// TIA Portal project "YDSLK_HMI_2023-05-10_08-26_V3_00T" (V15.1) (continued)
   "ST_HMI_Var_HMI_r64_DingZi_Zouche_ratio_KongDing_65_1" : LReal = PLC ST_HMI_Var.HMI_r64_DingZi_Zouche_ratio_KongDing_65_1 AT 10-30-00-01-00-21-84-00-4D-40, 1 s
   "ST_Calculation_Var_g_i16_Calculation_0_Status" : Int = PLC ST_Calculation_Var.g_i16_Calculation_0_Status AT 10-05-00-01-00-13-84-00-00-00, 1 s
   "ST_1TCP_g_myStructSend__lreal_20" : LReal = PLC ST_1TCP.g_myStructSend._lreal_20 AT 10-30-00-01-00-0D-84-01-30-40, 1 s
   "ST_1TCP_g_myStructSend__lreal_1" : LReal = PLC ST_1TCP.g_myStructSend._lreal_1 AT 10-30-00-01-00-0D-84-01-2B-80, 1 s
   "ST_HMI_Var_HMI_bo_ZouChe_Holding_Brake_Open" : Bool = PLC ST_HMI_Var.HMI_bo_ZouChe_Holding_Brake_Open AT 10-01-00-01-00-21-84-00-72-50, 1 s
   "ST_Real_Monitoring_HMI_r64_Real_QianShen_WuNian" : LReal = PLC ST_Real_Monitoring.HMI_r64_Real_QianShen_WuNian AT 10-30-00-01-00-2D-84-00-00-00, 1 s
   "ST_Real_Monitoring_HMI_r64Axis_ZouChe_Position_JiZhong_QianShen_Start" : LReal = PLC ST_Real_Monitoring.HMI_r64Axis_ZouChe_Position_JiZhong_QianShen_Start AT 10-30-00-01-00-2D-84-00-00-40, 1 s
   "ST_Real_Monitoring_HMI_r64_NianDu_JiZhong_QianShen_Start" : LReal = PLC ST_Real_Monitoring.HMI_r64_NianDu_JiZhong_QianShen_Start AT 10-30-00-01-00-2D-84-00-00-80, 1 s
   "ST_Real_Monitoring_HMI_r64Axis_ZouChe_Position_LuoLa_Stop" : LReal = PLC ST_Real_Monitoring.HMI_r64Axis_ZouChe_Position_LuoLa_Stop AT 10-30-00-01-00-2D-84-00-00-C0, 1 s
   "ST_Real_Monitoring_HMI_r64_NianDu_LuoLa_Stop" : LReal = PLC ST_Real_Monitoring.HMI_r64_NianDu_LuoLa_Stop AT 10-30-00-01-00-2D-84-00-01-00, 1 s
   "ST_Real_Monitoring_HMI_r64Axis_ZouChe_Position_YiNian_DaoDa" : LReal = PLC ST_Real_Monitoring.HMI_r64Axis_ZouChe_Position_YiNian_DaoDa AT 10-30-00-01-00-2D-84-00-01-40, 1 s
   "ST_Convert_ReadParameters_g_r64_SERVO_03_ZouChe_35_Motor_temperature_real" : LReal = PLC ST_Convert_ReadParameters.g_r64_SERVO_03_ZouChe_35_Motor_temperature_real AT 10-30-00-01-00-18-84-00-00-C0, 1 s
   "ST_Convert_ReadParameters_g_r64_SERVO_03_ZouChe_37_4_Power_unit_temperatures_Interior_of_power_unit_real" : LReal = PLC ST_Convert_ReadParameters.g_r64_SERVO_03_ZouChe_37_4_Power_unit_temperatures_Interior_of_power_unit_real AT 10-30-00-01-00-18-84-00-01-40, 1 s
   "ST_Convert_ReadParameters_g_r64_SERVO_04_ZhangLi_35_Motor_temperature_real" : LReal = PLC ST_Convert_ReadParameters.g_r64_SERVO_04_ZhangLi_35_Motor_temperature_real AT 10-30-00-01-00-18-84-00-03-00, 1 s
   "ST_Convert_ReadParameters_g_r64_SERVO_05_ChengXing_35_Motor_temperature_real" : LReal = PLC ST_Convert_ReadParameters.g_r64_SERVO_05_ChengXing_35_Motor_temperature_real AT 10-30-00-01-00-18-84-00-05-40, 1 s
   "ST_Convert_ReadParameters_g_r64_SERVO_06_GunTong_35_Motor_temperature_real" : LReal = PLC ST_Convert_ReadParameters.g_r64_SERVO_06_GunTong_35_Motor_temperature_real AT 10-30-00-01-00-18-84-00-07-80, 1 s
   "ST_Convert_ReadParameters_g_r64_SERVO_08_LuoLa_35_Motor_temperature_real" : LReal = PLC ST_Convert_ReadParameters.g_r64_SERVO_08_LuoLa_35_Motor_temperature_real AT 10-30-00-01-00-18-84-00-0C-00, 1 s
   "ST_Convert_ReadParameters_g_r64_SERVO_07_DingZi_35_Motor_temperature_real" : LReal = PLC ST_Convert_ReadParameters.g_r64_SERVO_07_DingZi_35_Motor_temperature_real AT 10-30-00-01-00-18-84-00-09-C0, 1 s
   "ST_Convert_ReadParameters_g_r64_SERVO_05_ChengXing_37_4_Power_unit_temperatures_Interior_of_power_unit_real" : LReal = PLC ST_Convert_ReadParameters.g_r64_SERVO_05_ChengXing_37_4_Power_unit_temperatures_Interior_of_power_unit_real AT 10-30-00-01-00-18-84-00-05-C0, 1 s
   "ST_Convert_ReadParameters_g_r64_SERVO_07_DingZi_37_4_Power_unit_temperatures_Interior_of_power_unit_real" : LReal = PLC ST_Convert_ReadParameters.g_r64_SERVO_07_DingZi_37_4_Power_unit_temperatures_Interior_of_power_unit_real AT 10-30-00-01-00-18-84-00-0A-40, 1 s
   "ST_Convert_ReadParameters_g_r64_SERVO_08_LuoLa_37_4_Power_unit_temperatures_Interior_of_power_unit_real" : LReal = PLC ST_Convert_ReadParameters.g_r64_SERVO_08_LuoLa_37_4_Power_unit_temperatures_Interior_of_power_unit_real AT 10-30-00-01-00-18-84-00-0C-80, 1 s

HMI tags "变量表_卷绕经验参数"
   "ST_Calculation_Var_1_ZhiShu_ARRAY_JR{3}" : LReal = PLC ST_Calculation_Var_1.ZhiShu_ARRAY_JR[3] AT 10-30-00-01-00-14-84-00-22-00, 1 s
   "ST_Calculation_Var_1_ZhiShu_ARRAY_JR{4}" : LReal = PLC ST_Calculation_Var_1.ZhiShu_ARRAY_JR[4] AT 10-30-00-01-00-14-84-00-22-40, 1 s
   "ST_Calculation_Var_1_ZhiShu_ARRAY_JR{5}" : LReal = PLC ST_Calculation_Var_1.ZhiShu_ARRAY_JR[5] AT 10-30-00-01-00-14-84-00-22-80, 1 s
   "ST_Calculation_Var_1_ZhiShu_ARRAY_JR{6}" : LReal = PLC ST_Calculation_Var_1.ZhiShu_ARRAY_JR[6] AT 10-30-00-01-00-14-84-00-22-C0, 1 s
   "ST_Calculation_Var_1_ZhiShu_ARRAY_JR{7}" : LReal = PLC ST_Calculation_Var_1.ZhiShu_ARRAY_JR[7] AT 10-30-00-01-00-14-84-00-23-00, 1 s
   "ST_Calculation_Var_1_ZhiShu_ARRAY_JR{8}" : LReal = PLC ST_Calculation_Var_1.ZhiShu_ARRAY_JR[8] AT 10-30-00-01-00-14-84-00-23-40, 1 s
   "ST_Calculation_Var_1_ZhiShu_ARRAY_JR{9}" : LReal = PLC ST_Calculation_Var_1.ZhiShu_ARRAY_JR[9] AT 10-30-00-01-00-14-84-00-23-80, 1 s
   "ST_Calculation_Var_1_ZhiShu_ARRAY_JR{10}" : LReal = PLC ST_Calculation_Var_1.ZhiShu_ARRAY_JR[10] AT 10-30-00-01-00-14-84-00-23-C0, 1 s
   "ST_Calculation_Var_1_ZhiShu_ARRAY_JR{11}" : LReal = PLC ST_Calculation_Var_1.ZhiShu_ARRAY_JR[11] AT 10-30-00-01-00-14-84-00-24-00, 1 s
   "ST_Calculation_Var_1_ZhiShu_ARRAY_JR{12}" : LReal = PLC ST_Calculation_Var_1.ZhiShu_ARRAY_JR[12] AT 10-30-00-01-00-14-84-00-24-40, 1 s
   "ST_Calculation_Var_1_ZhiShu_ARRAY_JR{13}" : LReal = PLC ST_Calculation_Var_1.ZhiShu_ARRAY_JR[13] AT 10-30-00-01-00-14-84-00-24-80, 1 s
   "ST_Calculation_Var_1_ZhiShu_ARRAY_JR{14}" : LReal = PLC ST_Calculation_Var_1.ZhiShu_ARRAY_JR[14] AT 10-30-00-01-00-14-84-00-24-C0, 1 s
   "ST_Calculation_Var_1_ZhiShu_ARRAY_JR{15}" : LReal = PLC ST_Calculation_Var_1.ZhiShu_ARRAY_JR[15] AT 10-30-00-01-00-14-84-00-25-00, 1 s
   "ST_Calculation_Var_1_ZhiShu_ARRAY_JR{16}" : LReal = PLC ST_Calculation_Var_1.ZhiShu_ARRAY_JR[16] AT 10-30-00-01-00-14-84-00-25-40, 1 s
   "ST_Calculation_Var_1_ZhiShu_ARRAY_JR{17}" : LReal = PLC ST_Calculation_Var_1.ZhiShu_ARRAY_JR[17] AT 10-30-00-01-00-14-84-00-25-80, 1 s
   "ST_Calculation_Var_1_ZhiShu_ARRAY_JR{18}" : LReal = PLC ST_Calculation_Var_1.ZhiShu_ARRAY_JR[18] AT 10-30-00-01-00-14-84-00-25-C0, 1 s
   "ST_Calculation_Var_1_ZhiShu_ARRAY_JR{19}" : LReal = PLC ST_Calculation_Var_1.ZhiShu_ARRAY_JR[19] AT 10-30-00-01-00-14-84-00-26-00, 1 s
   "ST_Calculation_Var_1_ZhiShu_ARRAY_JR{20}" : LReal = PLC ST_Calculation_Var_1.ZhiShu_ARRAY_JR[20] AT 10-30-00-01-00-14-84-00-26-40, 1 s
   "ST_Calculation_Var_1_ZhiShu_ARRAY_JR{21}" : LReal = PLC ST_Calculation_Var_1.ZhiShu_ARRAY_JR[21] AT 10-30-00-01-00-14-84-00-26-80, 1 s
   "ST_Calculation_Var_1_ZhiShu_ARRAY_JR{22}" : LReal = PLC ST_Calculation_Var_1.ZhiShu_ARRAY_JR[22] AT 10-30-00-01-00-14-84-00-26-C0, 1 s
   "ST_Calculation_Var_1_ZhiShu_ARRAY_JR{23}" : LReal = PLC ST_Calculation_Var_1.ZhiShu_ARRAY_JR[23] AT 10-30-00-01-00-14-84-00-27-00, 1 s
   "ST_Calculation_Var_1_ZhiShu_ARRAY_JR{24}" : LReal = PLC ST_Calculation_Var_1.ZhiShu_ARRAY_JR[24] AT 10-30-00-01-00-14-84-00-27-40, 1 s
   "ST_Calculation_Var_1_ZhiShu_ARRAY_JR{25}" : LReal = PLC ST_Calculation_Var_1.ZhiShu_ARRAY_JR[25] AT 10-30-00-01-00-14-84-00-27-80, 1 s
   "ST_Calculation_Var_1_ZhiShu_ARRAY_JR{26}" : LReal = PLC ST_Calculation_Var_1.ZhiShu_ARRAY_JR[26] AT 10-30-00-01-00-14-84-00-27-C0, 1 s
   "ST_Calculation_Var_1_ZhiShu_ARRAY_JR{27}" : LReal = PLC ST_Calculation_Var_1.ZhiShu_ARRAY_JR[27] AT 10-30-00-01-00-14-84-00-28-00, 1 s
   "ST_Calculation_Var_1_ZhiShu_ARRAY_JR{28}" : LReal = PLC ST_Calculation_Var_1.ZhiShu_ARRAY_JR[28] AT 10-30-00-01-00-14-84-00-28-40, 1 s
   "ST_Calculation_Var_1_ZhiShu_ARRAY_JR{29}" : LReal = PLC ST_Calculation_Var_1.ZhiShu_ARRAY_JR[29] AT 10-30-00-01-00-14-84-00-28-80, 1 s
   "ST_Calculation_Var_1_ZhiShu_ARRAY_JR{30}" : LReal = PLC ST_Calculation_Var_1.ZhiShu_ARRAY_JR[30] AT 10-30-00-01-00-14-84-00-28-C0, 1 s
   "ST_Calculation_Var_1_ZhiShu_ARRAY_JR{31}" : LReal = PLC ST_Calculation_Var_1.ZhiShu_ARRAY_JR[31] AT 10-30-00-01-00-14-84-00-29-00, 1 s
   "ST_Calculation_Var_1_ZhiShu_ARRAY_JR{32}" : LReal = PLC ST_Calculation_Var_1.ZhiShu_ARRAY_JR[32] AT 10-30-00-01-00-14-84-00-29-40, 1 s
   "ST_Calculation_Var_1_ZhiShu_ARRAY_JR{33}" : LReal = PLC ST_Calculation_Var_1.ZhiShu_ARRAY_JR[33] AT 10-30-00-01-00-14-84-00-29-80, 1 s
   "ST_Calculation_Var_1_ZhiShu_ARRAY_JR{34}" : LReal = PLC ST_Calculation_Var_1.ZhiShu_ARRAY_JR[34] AT 10-30-00-01-00-14-84-00-29-C0, 1 s
   "ST_Calculation_Var_1_ZhiShu_ARRAY_JR{35}" : LReal = PLC ST_Calculation_Var_1.ZhiShu_ARRAY_JR[35] AT 10-30-00-01-00-14-84-00-2A-00, 1 s
   "ST_Calculation_Var_1_ZhiShu_ARRAY_JR{36}" : LReal = PLC ST_Calculation_Var_1.ZhiShu_ARRAY_JR[36] AT 10-30-00-01-00-14-84-00-2A-40, 1 s
   "ST_Calculation_Var_1_ZhiShu_ARRAY_JR{37}" : LReal = PLC ST_Calculation_Var_1.ZhiShu_ARRAY_JR[37] AT 10-30-00-01-00-14-84-00-2A-80, 1 s
   "ST_Calculation_Var_1_ZhiShu_ARRAY_JR{38}" : LReal = PLC ST_Calculation_Var_1.ZhiShu_ARRAY_JR[38] AT 10-30-00-01-00-14-84-00-2A-C0, 1 s
   "ST_Calculation_Var_1_ZhiShu_ARRAY_JR{39}" : LReal = PLC ST_Calculation_Var_1.ZhiShu_ARRAY_JR[39] AT 10-30-00-01-00-14-84-00-2B-00, 1 s
   "ST_Calculation_Var_1_ZhiShu_ARRAY_JR{40}" : LReal = PLC ST_Calculation_Var_1.ZhiShu_ARRAY_JR[40] AT 10-30-00-01-00-14-84-00-2B-40, 1 s
   "ST_Calculation_Var_1_ZhiShu_ARRAY_JR{41}" : LReal = PLC ST_Calculation_Var_1.ZhiShu_ARRAY_JR[41] AT 10-30-00-01-00-14-84-00-2B-80, 1 s
   "ST_Calculation_Var_1_ZhiShu_ARRAY_JR{42}" : LReal = PLC ST_Calculation_Var_1.ZhiShu_ARRAY_JR[42] AT 10-30-00-01-00-14-84-00-2B-C0, 1 s
   "ST_Calculation_Var_1_ZhiShu_ARRAY_JR{43}" : LReal = PLC ST_Calculation_Var_1.ZhiShu_ARRAY_JR[43] AT 10-30-00-01-00-14-84-00-2C-00, 1 s
   "ST_Calculation_Var_1_ZhiShu_ARRAY_JR{44}" : LReal = PLC ST_Calculation_Var_1.ZhiShu_ARRAY_JR[44] AT 10-30-00-01-00-14-84-00-2C-40, 1 s
   "ST_Calculation_Var_1_ZhiShu_ARRAY_JR{45}" : LReal = PLC ST_Calculation_Var_1.ZhiShu_ARRAY_JR[45] AT 10-30-00-01-00-14-84-00-2C-80, 1 s
   "ST_Calculation_Var_1_ZhiShu_ARRAY_JR{46}" : LReal = PLC ST_Calculation_Var_1.ZhiShu_ARRAY_JR[46] AT 10-30-00-01-00-14-84-00-2C-C0, 1 s
   "ST_Calculation_Var_1_ZhiShu_ARRAY_JR{47}" : LReal = PLC ST_Calculation_Var_1.ZhiShu_ARRAY_JR[47] AT 10-30-00-01-00-14-84-00-2D-00, 1 s
   "ST_Calculation_Var_1_f1_n_delt_0_n_ARRAY_JR{3}" : LReal = PLC ST_Calculation_Var_1.f1_n_delt_0_n_ARRAY_JR[3] AT 10-30-00-01-00-14-84-00-2E-00, 1 s
   "ST_Calculation_Var_1_f1_n_delt_0_n_ARRAY_JR{4}" : LReal = PLC ST_Calculation_Var_1.f1_n_delt_0_n_ARRAY_JR[4] AT 10-30-00-01-00-14-84-00-2E-40, 1 s
   "ST_Calculation_Var_1_f1_n_delt_0_n_ARRAY_JR{5}" : LReal = PLC ST_Calculation_Var_1.f1_n_delt_0_n_ARRAY_JR[5] AT 10-30-00-01-00-14-84-00-2E-80, 1 s
   "ST_Calculation_Var_1_f1_n_delt_0_n_ARRAY_JR{6}" : LReal = PLC ST_Calculation_Var_1.f1_n_delt_0_n_ARRAY_JR[6] AT 10-30-00-01-00-14-84-00-2E-C0, 1 s
   "ST_Calculation_Var_1_f1_n_delt_0_n_ARRAY_JR{7}" : LReal = PLC ST_Calculation_Var_1.f1_n_delt_0_n_ARRAY_JR[7] AT 10-30-00-01-00-14-84-00-2F-00, 1 s
   "ST_Calculation_Var_1_f1_n_delt_0_n_ARRAY_JR{8}" : LReal = PLC ST_Calculation_Var_1.f1_n_delt_0_n_ARRAY_JR[8] AT 10-30-00-01-00-14-84-00-2F-40, 1 s
   "ST_Calculation_Var_1_f1_n_delt_0_n_ARRAY_JR{9}" : LReal = PLC ST_Calculation_Var_1.f1_n_delt_0_n_ARRAY_JR[9] AT 10-30-00-01-00-14-84-00-2F-80, 1 s
   "ST_Calculation_Var_1_f1_n_delt_0_n_ARRAY_JR{10}" : LReal = PLC ST_Calculation_Var_1.f1_n_delt_0_n_ARRAY_JR[10] AT 10-30-00-01-00-14-84-00-2F-C0, 1 s
   "ST_Calculation_Var_1_f1_n_delt_0_n_ARRAY_JR{11}" : LReal = PLC ST_Calculation_Var_1.f1_n_delt_0_n_ARRAY_JR[11] AT 10-30-00-01-00-14-84-00-30-00, 1 s
   "ST_Calculation_Var_1_f1_n_delt_0_n_ARRAY_JR{12}" : LReal = PLC ST_Calculation_Var_1.f1_n_delt_0_n_ARRAY_JR[12] AT 10-30-00-01-00-14-84-00-30-40, 1 s
   "ST_Calculation_Var_1_f1_n_delt_0_n_ARRAY_JR{13}" : LReal = PLC ST_Calculation_Var_1.f1_n_delt_0_n_ARRAY_JR[13] AT 10-30-00-01-00-14-84-00-30-80, 1 s
   "ST_Calculation_Var_1_f1_n_delt_0_n_ARRAY_JR{14}" : LReal = PLC ST_Calculation_Var_1.f1_n_delt_0_n_ARRAY_JR[14] AT 10-30-00-01-00-14-84-00-30-C0, 1 s
   "ST_Calculation_Var_1_f1_n_delt_0_n_ARRAY_JR{15}" : LReal = PLC ST_Calculation_Var_1.f1_n_delt_0_n_ARRAY_JR[15] AT 10-30-00-01-00-14-84-00-31-00, 1 s
   "ST_Calculation_Var_1_f1_n_delt_0_n_ARRAY_JR{16}" : LReal = PLC ST_Calculation_Var_1.f1_n_delt_0_n_ARRAY_JR[16] AT 10-30-00-01-00-14-84-00-31-40, 1 s
   "ST_Calculation_Var_1_f1_n_delt_0_n_ARRAY_JR{17}" : LReal = PLC ST_Calculation_Var_1.f1_n_delt_0_n_ARRAY_JR[17] AT 10-30-00-01-00-14-84-00-31-80, 1 s
   "ST_Calculation_Var_1_f1_n_delt_0_n_ARRAY_JR{18}" : LReal = PLC ST_Calculation_Var_1.f1_n_delt_0_n_ARRAY_JR[18] AT 10-30-00-01-00-14-84-00-31-C0, 1 s
   "ST_Calculation_Var_1_f1_n_delt_0_n_ARRAY_JR{19}" : LReal = PLC ST_Calculation_Var_1.f1_n_delt_0_n_ARRAY_JR[19] AT 10-30-00-01-00-14-84-00-32-00, 1 s
   "ST_Calculation_Var_1_f1_n_delt_0_n_ARRAY_JR{20}" : LReal = PLC ST_Calculation_Var_1.f1_n_delt_0_n_ARRAY_JR[20] AT 10-30-00-01-00-14-84-00-32-40, 1 s
   "ST_Calculation_Var_1_f1_n_delt_0_n_ARRAY_JR{21}" : LReal = PLC ST_Calculation_Var_1.f1_n_delt_0_n_ARRAY_JR[21] AT 10-30-00-01-00-14-84-00-32-80, 1 s
   "ST_Calculation_Var_1_f1_n_delt_0_n_ARRAY_JR{22}" : LReal = PLC ST_Calculation_Var_1.f1_n_delt_0_n_ARRAY_JR[22] AT 10-30-00-01-00-14-84-00-32-C0, 1 s
   "ST_Calculation_Var_1_f1_n_delt_0_n_ARRAY_JR{23}" : LReal = PLC ST_Calculation_Var_1.f1_n_delt_0_n_ARRAY_JR[23] AT 10-30-00-01-00-14-84-00-33-00, 1 s
   "ST_Calculation_Var_1_f1_n_delt_0_n_ARRAY_JR{24}" : LReal = PLC ST_Calculation_Var_1.f1_n_delt_0_n_ARRAY_JR[24] AT 10-30-00-01-00-14-84-00-33-40, 1 s
   "ST_Calculation_Var_1_f1_n_delt_0_n_ARRAY_JR{25}" : LReal = PLC ST_Calculation_Var_1.f1_n_delt_0_n_ARRAY_JR[25] AT 10-30-00-01-00-14-84-00-33-80, 1 s
   "ST_Calculation_Var_1_f1_n_delt_0_n_ARRAY_JR{26}" : LReal = PLC ST_Calculation_Var_1.f1_n_delt_0_n_ARRAY_JR[26] AT 10-30-00-01-00-14-84-00-33-C0, 1 s
   "ST_Calculation_Var_1_f1_n_delt_0_n_ARRAY_JR{27}" : LReal = PLC ST_Calculation_Var_1.f1_n_delt_0_n_ARRAY_JR[27] AT 10-30-00-01-00-14-84-00-34-00, 1 s
   "ST_Calculation_Var_1_f1_n_delt_0_n_ARRAY_JR{28}" : LReal = PLC ST_Calculation_Var_1.f1_n_delt_0_n_ARRAY_JR[28] AT 10-30-00-01-00-14-84-00-34-40, 1 s
   "ST_Calculation_Var_1_f1_n_delt_0_n_ARRAY_JR{29}" : LReal = PLC ST_Calculation_Var_1.f1_n_delt_0_n_ARRAY_JR[29] AT 10-30-00-01-00-14-84-00-34-80, 1 s
   "ST_Calculation_Var_1_f1_n_delt_0_n_ARRAY_JR{30}" : LReal = PLC ST_Calculation_Var_1.f1_n_delt_0_n_ARRAY_JR[30] AT 10-30-00-01-00-14-84-00-34-C0, 1 s
   "ST_Calculation_Var_1_f1_n_delt_0_n_ARRAY_JR{31}" : LReal = PLC ST_Calculation_Var_1.f1_n_delt_0_n_ARRAY_JR[31] AT 10-30-00-01-00-14-84-00-35-00, 1 s
   "ST_Calculation_Var_1_f1_n_delt_0_n_ARRAY_JR{32}" : LReal = PLC ST_Calculation_Var_1.f1_n_delt_0_n_ARRAY_JR[32] AT 10-30-00-01-00-14-84-00-35-40, 1 s
   "ST_Calculation_Var_1_f1_n_delt_0_n_ARRAY_JR{33}" : LReal = PLC ST_Calculation_Var_1.f1_n_delt_0_n_ARRAY_JR[33] AT 10-30-00-01-00-14-84-00-35-80, 1 s
   "ST_Calculation_Var_1_f1_n_delt_0_n_ARRAY_JR{34}" : LReal = PLC ST_Calculation_Var_1.f1_n_delt_0_n_ARRAY_JR[34] AT 10-30-00-01-00-14-84-00-35-C0, 1 s
   "ST_Calculation_Var_1_f1_n_delt_0_n_ARRAY_JR{35}" : LReal = PLC ST_Calculation_Var_1.f1_n_delt_0_n_ARRAY_JR[35] AT 10-30-00-01-00-14-84-00-36-00, 1 s
   "ST_Calculation_Var_1_f1_n_delt_0_n_ARRAY_JR{36}" : LReal = PLC ST_Calculation_Var_1.f1_n_delt_0_n_ARRAY_JR[36] AT 10-30-00-01-00-14-84-00-36-40, 1 s
   "ST_Calculation_Var_1_f1_n_delt_0_n_ARRAY_JR{37}" : LReal = PLC ST_Calculation_Var_1.f1_n_delt_0_n_ARRAY_JR[37] AT 10-30-00-01-00-14-84-00-36-80, 1 s
   "ST_Calculation_Var_1_f1_n_delt_0_n_ARRAY_JR{38}" : LReal = PLC ST_Calculation_Var_1.f1_n_delt_0_n_ARRAY_JR[38] AT 10-30-00-01-00-14-84-00-36-C0, 1 s
   "ST_Calculation_Var_1_f1_n_delt_0_n_ARRAY_JR{39}" : LReal = PLC ST_Calculation_Var_1.f1_n_delt_0_n_ARRAY_JR[39] AT 10-30-00-01-00-14-84-00-37-00, 1 s
   "ST_Calculation_Var_1_f1_n_delt_0_n_ARRAY_JR{40}" : LReal = PLC ST_Calculation_Var_1.f1_n_delt_0_n_ARRAY_JR[40] AT 10-30-00-01-00-14-84-00-37-40, 1 s
   "ST_Calculation_Var_1_f1_n_delt_0_n_ARRAY_JR{41}" : LReal = PLC ST_Calculation_Var_1.f1_n_delt_0_n_ARRAY_JR[41] AT 10-30-00-01-00-14-84-00-37-80, 1 s
   "ST_Calculation_Var_1_f1_n_delt_0_n_ARRAY_JR{42}" : LReal = PLC ST_Calculation_Var_1.f1_n_delt_0_n_ARRAY_JR[42] AT 10-30-00-01-00-14-84-00-37-C0, 1 s
   "ST_Calculation_Var_1_f1_n_delt_0_n_ARRAY_JR{43}" : LReal = PLC ST_Calculation_Var_1.f1_n_delt_0_n_ARRAY_JR[43] AT 10-30-00-01-00-14-84-00-38-00, 1 s
   "ST_Calculation_Var_1_f1_n_delt_0_n_ARRAY_JR{44}" : LReal = PLC ST_Calculation_Var_1.f1_n_delt_0_n_ARRAY_JR[44] AT 10-30-00-01-00-14-84-00-38-40, 1 s
   "ST_Calculation_Var_1_f1_n_delt_0_n_ARRAY_JR{45}" : LReal = PLC ST_Calculation_Var_1.f1_n_delt_0_n_ARRAY_JR[45] AT 10-30-00-01-00-14-84-00-38-80, 1 s
   "ST_Calculation_Var_1_f1_n_delt_0_n_ARRAY_JR{46}" : LReal = PLC ST_Calculation_Var_1.f1_n_delt_0_n_ARRAY_JR[46] AT 10-30-00-01-00-14-84-00-38-C0, 1 s
   "ST_Calculation_Var_1_f1_n_delt_0_n_ARRAY_JR{47}" : LReal = PLC ST_Calculation_Var_1.f1_n_delt_0_n_ARRAY_JR[47] AT 10-30-00-01-00-14-84-00-39-00, 1 s
   "ST_Calculation_Var_1_g1_n_delt_0_n_ARRAY_JR{3}" : LReal = PLC ST_Calculation_Var_1.g1_n_delt_0_n_ARRAY_JR[3] AT 10-30-00-01-00-14-84-00-3A-00, 1 s
   "ST_Calculation_Var_1_g1_n_delt_0_n_ARRAY_JR{4}" : LReal = PLC ST_Calculation_Var_1.g1_n_delt_0_n_ARRAY_JR[4] AT 10-30-00-01-00-14-84-00-3A-40, 1 s
   "ST_Calculation_Var_1_g1_n_delt_0_n_ARRAY_JR{5}" : LReal = PLC ST_Calculation_Var_1.g1_n_delt_0_n_ARRAY_JR[5] AT 10-30-00-01-00-14-84-00-3A-80, 1 s
   "ST_Calculation_Var_1_g1_n_delt_0_n_ARRAY_JR{6}" : LReal = PLC ST_Calculation_Var_1.g1_n_delt_0_n_ARRAY_JR[6] AT 10-30-00-01-00-14-84-00-3A-C0, 1 s
   "ST_Calculation_Var_1_g1_n_delt_0_n_ARRAY_JR{7}" : LReal = PLC ST_Calculation_Var_1.g1_n_delt_0_n_ARRAY_JR[7] AT 10-30-00-01-00-14-84-00-3B-00, 1 s
   "ST_Calculation_Var_1_g1_n_delt_0_n_ARRAY_JR{8}" : LReal = PLC ST_Calculation_Var_1.g1_n_delt_0_n_ARRAY_JR[8] AT 10-30-00-01-00-14-84-00-3B-40, 1 s
   "ST_Calculation_Var_1_g1_n_delt_0_n_ARRAY_JR{9}" : LReal = PLC ST_Calculation_Var_1.g1_n_delt_0_n_ARRAY_JR[9] AT 10-30-00-01-00-14-84-00-3B-80, 1 s
   "ST_Calculation_Var_1_g1_n_delt_0_n_ARRAY_JR{10}" : LReal = PLC ST_Calculation_Var_1.g1_n_delt_0_n_ARRAY_JR[10] AT 10-30-00-01-00-14-84-00-3B-C0, 1 s
   "ST_Calculation_Var_1_g1_n_delt_0_n_ARRAY_JR{11}" : LReal = PLC ST_Calculation_Var_1.g1_n_delt_0_n_ARRAY_JR[11] AT 10-30-00-01-00-14-84-00-3C-00, 1 s
   "ST_Calculation_Var_1_g1_n_delt_0_n_ARRAY_JR{12}" : LReal = PLC ST_Calculation_Var_1.g1_n_delt_0_n_ARRAY_JR[12] AT 10-30-00-01-00-14-84-00-3C-40, 1 s
   "ST_Calculation_Var_1_g1_n_delt_0_n_ARRAY_JR{13}" : LReal = PLC ST_Calculation_Var_1.g1_n_delt_0_n_ARRAY_JR[13] AT 10-30-00-01-00-14-84-00-3C-80, 1 s
   "ST_Calculation_Var_1_g1_n_delt_0_n_ARRAY_JR{14}" : LReal = PLC ST_Calculation_Var_1.g1_n_delt_0_n_ARRAY_JR[14] AT 10-30-00-01-00-14-84-00-3C-C0, 1 s
   "ST_Calculation_Var_1_g1_n_delt_0_n_ARRAY_JR{15}" : LReal = PLC ST_Calculation_Var_1.g1_n_delt_0_n_ARRAY_JR[15] AT 10-30-00-01-00-14-84-00-3D-00, 1 s
   "ST_Calculation_Var_1_g1_n_delt_0_n_ARRAY_JR{16}" : LReal = PLC ST_Calculation_Var_1.g1_n_delt_0_n_ARRAY_JR[16] AT 10-30-00-01-00-14-84-00-3D-40, 1 s
   "ST_Calculation_Var_1_g1_n_delt_0_n_ARRAY_JR{17}" : LReal = PLC ST_Calculation_Var_1.g1_n_delt_0_n_ARRAY_JR[17] AT 10-30-00-01-00-14-84-00-3D-80, 1 s
   "ST_Calculation_Var_1_g1_n_delt_0_n_ARRAY_JR{18}" : LReal = PLC ST_Calculation_Var_1.g1_n_delt_0_n_ARRAY_JR[18] AT 10-30-00-01-00-14-84-00-3D-C0, 1 s
   "ST_Calculation_Var_1_g1_n_delt_0_n_ARRAY_JR{19}" : LReal = PLC ST_Calculation_Var_1.g1_n_delt_0_n_ARRAY_JR[19] AT 10-30-00-01-00-14-84-00-3E-00, 1 s
   "ST_Calculation_Var_1_g1_n_delt_0_n_ARRAY_JR{20}" : LReal = PLC ST_Calculation_Var_1.g1_n_delt_0_n_ARRAY_JR[20] AT 10-30-00-01-00-14-84-00-3E-40, 1 s
   "ST_Calculation_Var_1_g1_n_delt_0_n_ARRAY_JR{21}" : LReal = PLC ST_Calculation_Var_1.g1_n_delt_0_n_ARRAY_JR[21] AT 10-30-00-01-00-14-84-00-3E-80, 1 s
   "ST_Calculation_Var_1_g1_n_delt_0_n_ARRAY_JR{22}" : LReal = PLC ST_Calculation_Var_1.g1_n_delt_0_n_ARRAY_JR[22] AT 10-30-00-01-00-14-84-00-3E-C0, 1 s
   "ST_Calculation_Var_1_g1_n_delt_0_n_ARRAY_JR{23}" : LReal = PLC ST_Calculation_Var_1.g1_n_delt_0_n_ARRAY_JR[23] AT 10-30-00-01-00-14-84-00-3F-00, 1 s
   "ST_Calculation_Var_1_g1_n_delt_0_n_ARRAY_JR{24}" : LReal = PLC ST_Calculation_Var_1.g1_n_delt_0_n_ARRAY_JR[24] AT 10-30-00-01-00-14-84-00-3F-40, 1 s
   "ST_Calculation_Var_1_g1_n_delt_0_n_ARRAY_JR{25}" : LReal = PLC ST_Calculation_Var_1.g1_n_delt_0_n_ARRAY_JR[25] AT 10-30-00-01-00-14-84-00-3F-80, 1 s
   "ST_Calculation_Var_1_g1_n_delt_0_n_ARRAY_JR{26}" : LReal = PLC ST_Calculation_Var_1.g1_n_delt_0_n_ARRAY_JR[26] AT 10-30-00-01-00-14-84-00-3F-C0, 1 s
   "ST_Calculation_Var_1_g1_n_delt_0_n_ARRAY_JR{27}" : LReal = PLC ST_Calculation_Var_1.g1_n_delt_0_n_ARRAY_JR[27] AT 10-30-00-01-00-14-84-00-40-00, 1 s
   "ST_Calculation_Var_1_g1_n_delt_0_n_ARRAY_JR{28}" : LReal = PLC ST_Calculation_Var_1.g1_n_delt_0_n_ARRAY_JR[28] AT 10-30-00-01-00-14-84-00-40-40, 1 s
   "ST_Calculation_Var_1_g1_n_delt_0_n_ARRAY_JR{29}" : LReal = PLC ST_Calculation_Var_1.g1_n_delt_0_n_ARRAY_JR[29] AT 10-30-00-01-00-14-84-00-40-80, 1 s
   "ST_Calculation_Var_1_g1_n_delt_0_n_ARRAY_JR{30}" : LReal = PLC ST_Calculation_Var_1.g1_n_delt_0_n_ARRAY_JR[30] AT 10-30-00-01-00-14-84-00-40-C0, 1 s
   "ST_Calculation_Var_1_g1_n_delt_0_n_ARRAY_JR{31}" : LReal = PLC ST_Calculation_Var_1.g1_n_delt_0_n_ARRAY_JR[31] AT 10-30-00-01-00-14-84-00-41-00, 1 s
   "ST_Calculation_Var_1_g1_n_delt_0_n_ARRAY_JR{32}" : LReal = PLC ST_Calculation_Var_1.g1_n_delt_0_n_ARRAY_JR[32] AT 10-30-00-01-00-14-84-00-41-40, 1 s
   "ST_Calculation_Var_1_g1_n_delt_0_n_ARRAY_JR{33}" : LReal = PLC ST_Calculation_Var_1.g1_n_delt_0_n_ARRAY_JR[33] AT 10-30-00-01-00-14-84-00-41-80, 1 s
   "ST_Calculation_Var_1_g1_n_delt_0_n_ARRAY_JR{34}" : LReal = PLC ST_Calculation_Var_1.g1_n_delt_0_n_ARRAY_JR[34] AT 10-30-00-01-00-14-84-00-41-C0, 1 s
   "ST_Calculation_Var_1_g1_n_delt_0_n_ARRAY_JR{35}" : LReal = PLC ST_Calculation_Var_1.g1_n_delt_0_n_ARRAY_JR[35] AT 10-30-00-01-00-14-84-00-42-00, 1 s
   "ST_Calculation_Var_1_g1_n_delt_0_n_ARRAY_JR{36}" : LReal = PLC ST_Calculation_Var_1.g1_n_delt_0_n_ARRAY_JR[36] AT 10-30-00-01-00-14-84-00-42-40, 1 s
   "ST_Calculation_Var_1_g1_n_delt_0_n_ARRAY_JR{37}" : LReal = PLC ST_Calculation_Var_1.g1_n_delt_0_n_ARRAY_JR[37] AT 10-30-00-01-00-14-84-00-42-80, 1 s
   "ST_Calculation_Var_1_g1_n_delt_0_n_ARRAY_JR{38}" : LReal = PLC ST_Calculation_Var_1.g1_n_delt_0_n_ARRAY_JR[38] AT 10-30-00-01-00-14-84-00-42-C0, 1 s
   "ST_Calculation_Var_1_g1_n_delt_0_n_ARRAY_JR{39}" : LReal = PLC ST_Calculation_Var_1.g1_n_delt_0_n_ARRAY_JR[39] AT 10-30-00-01-00-14-84-00-43-00, 1 s
   "ST_Calculation_Var_1_g1_n_delt_0_n_ARRAY_JR{40}" : LReal = PLC ST_Calculation_Var_1.g1_n_delt_0_n_ARRAY_JR[40] AT 10-30-00-01-00-14-84-00-43-40, 1 s
   "ST_Calculation_Var_1_g1_n_delt_0_n_ARRAY_JR{41}" : LReal = PLC ST_Calculation_Var_1.g1_n_delt_0_n_ARRAY_JR[41] AT 10-30-00-01-00-14-84-00-43-80, 1 s
   "ST_Calculation_Var_1_g1_n_delt_0_n_ARRAY_JR{42}" : LReal = PLC ST_Calculation_Var_1.g1_n_delt_0_n_ARRAY_JR[42] AT 10-30-00-01-00-14-84-00-43-C0, 1 s
   "ST_Calculation_Var_1_g1_n_delt_0_n_ARRAY_JR{43}" : LReal = PLC ST_Calculation_Var_1.g1_n_delt_0_n_ARRAY_JR[43] AT 10-30-00-01-00-14-84-00-44-00, 1 s
   "ST_Calculation_Var_1_g1_n_delt_0_n_ARRAY_JR{44}" : LReal = PLC ST_Calculation_Var_1.g1_n_delt_0_n_ARRAY_JR[44] AT 10-30-00-01-00-14-84-00-44-40, 1 s
   "ST_Calculation_Var_1_g1_n_delt_0_n_ARRAY_JR{45}" : LReal = PLC ST_Calculation_Var_1.g1_n_delt_0_n_ARRAY_JR[45] AT 10-30-00-01-00-14-84-00-44-80, 1 s
   "ST_Calculation_Var_1_g1_n_delt_0_n_ARRAY_JR{46}" : LReal = PLC ST_Calculation_Var_1.g1_n_delt_0_n_ARRAY_JR[46] AT 10-30-00-01-00-14-84-00-44-C0, 1 s
   "ST_Calculation_Var_1_g1_n_delt_0_n_ARRAY_JR{47}" : LReal = PLC ST_Calculation_Var_1.g1_n_delt_0_n_ARRAY_JR[47] AT 10-30-00-01-00-14-84-00-45-00, 1 s

text list "Text list_MasterMode": 1 'ABSOLUTE'; 45 'EFFECTIVE'; 115 'RELATIVE'; 149 'USER_DEFAULT'

text list "mode_enabled_2": 1 '故障中 / Error / 고장중'; 2 '无使能 / Disable / 무능력'; 4 '手动 / Manual / 手動 / 수동'; 8 '定位中 / Startposition / 위치유도'; 16 '管前生头 / Atuomatic / pipe front 스레딩'; 32 '管后生头 / NothingSelect / pipe rear 스레딩'; 64 '自动 / Changing / 自動 / 자동'; 128 '没选择 / 선택하지 않았음'

text list "Text list_mergeMode": 60 'IMMEDIATELY'; 89 'NEXT_MOTION'; 119 'SEQUENTIAL'; 142 'SUPERIMPOSED_MOTION_MERGE'

text list "Text list_negativeAccelEndJerkType": 40 'DIRECT'; 45 'EFFECTIVE'; 149 'USER_DEFAULT'

text list "Text list_negativeAccelStartJerkType": 40 'DIRECT'; 45 'EFFECTIVE'; 149 'USER_DEFAULT'

text list "Text list_positiveAccelEndJerkType": 40 'DIRECT'; 45 'EFFECTIVE'; 149 'USER_DEFAULT'

text list "mode_enabled": 1 'Mode:Error'; 2 'Mode:Disable'; 4 'Mode:Manual'; 8 'Mode:StartPosition'; 16 'Mode:KongDing / Mode:Automatic'; 32 'Mode:LuoSha / Mode:NothingSelected'; 64 'Mode:Automatic / Mode:Changing'; 128 'Mode:NothingSelect'

text list "Text list_syncProfileReference": 45 'EFFECTIVE'; 113 'RELATE_SYNC_PROFILE_TO_LEADING_VALUE'; 114 'RELATE_SYNC_PROFILE_TO_TIME'; 149 'USER_DEFAULT'

text list "automatic_status": 1 'Auto Status:Waiting'; 2 'Auto Status:EmergeStop / Auto Status:MergeStop'; 4 'Auto Status:AtuoStop'; 8 'Auto Status:ChuChe'; 16 'Auto Status:ChuCheDao'; 32 'Auto Status:TuiRao'; 64 'Auto Status:JuanRao'; 128 'Auto Status:CunRao'

text list "Text list_synchronizingmode": 14 'AT_THE_END_OF_CAM_CYCLE'; 45 'EFFECTIVE'; 60 'IMMEDIATELY'; 90 'NEXT_WITH_REFERENCE'; 99 'ON_MASTER_AND_SLAVE_POSITION'; 100 'ON_MASTER_POSITION'; 149 'USER_DEFAULT'; 315 'IMMEDIATELY_AND_SLAVE_POSITION'

text list "Text list_positiveAccelYype": 40 'DIRECT'; 45 'EFFECTIVE'; 149 'USER_DEFAULT'

text list "Text list_positioningMode": 1 'ABSOLUTE'; 115 'RELATIVE'

text list "Text list_velocityProfile": 45 'EFFECTIVE'; 103 'PARABOLIC'; 122 'SINUSOIDAL'; 124 'SMOOTH'; 146 'TRAPEZOIDAL'; 149 'USER_DEFAULT'

text list "Text list_nextCommand": 12 'AT_DECELERATION_START'; 13 'AT_MOTION_START'; 60 'IMMEDIATELY'; 156 'WHEN_ACCELERATION_DONE'; 159 'WHEN_BUFFER_READY'; 162 'WHEN_INTERPOLATION_DONE'; 163 'WHEN_MOTION_DONE'

text list "Text list_syncOffPositionReference": 15 'AXIS_STOPPED_AT_POSITION'; 18 'BEGIN_TO_STOP_WHEN_POSITION_REACHED'; 45 'EFFECTIVE'; 137 'STOP_SYMMETRIC_WITH_POSITION'; 149 'USER_DEFAULT'

text list "automatic_status_2": 1 '等待 / Waiting / 待機 / 대기'; 2 '紧急停止 / MergeStop / 緊急停止 / 비상정지'; 4 '自动停止 / AtuoStop / 自動停止 / 자동 정지'; 8 '出车 / ChuChe / 出機 / 외진'; 16 '出车到 / ChuCheDao / 出機完了 / 외진도착'; 32 '退绕 / TuiRao / パッキングオフ / 언와인딩'; 64 '卷绕 / JuanRao / 巻取 / 와인딩'; 128 '存绕 / CunRao / 逆巻取 / 와인딩 저장'

text list "luosha_status#mig1": 0 '状态;等待中 / 상태: 대기중'; 1 '进程1:成形弓至锭底 / 프로세스 1: 성형보우(성형호랑)에서 스핀들 밑부분까지'; 2 '进程2:至锭底后卷绕 / 프로세스 2: 스핀들 밑부분까지 한후 와인딩'; 4 '进程3:成形弓至卷绕点 / 프로세스 3: 성형보우(성형호랑)에서 와인딩 포인트까지'; 8 '进程4:放开张力弓 / 프로세스 4: 장력보우(장력호랑)를 풀기'; 16 '进程5:调整张力弓高低 / 프로세스 5: 장력보우(장력호랑) 높낮이를 조절'; 32 '状态:进行中1 / 상태: 진행중1'; 64 '状态:暂停中 / 상태: 일시 정지중'; 128 '状态:进行中2 / 상태: 진행중2'; 256 '进程9:存绕 / 프로세스 9: 와인딩 저장'

text list "Pictures": 1 '开始画面'; 2 '设置画面'; 3 '手动画面 / 手動画面 / 수동화면'; 4 '自动画面 / 自動画面 / 자동화면'; 5 '时间显示画面'; 6 '报警画面'; 7 '调试画面'; 8 '帮助画面'; 9 '用户管理画面'; 10 '工艺设置画面'; 12 '生头画面'; 13 '生头画面'; 21 '生头工艺设置画面'; 31 '工艺设置画面'; 38 '保养提示画面'

text list "Text list_movingMode": 180 'POSITION_CONTROLLED'; 181 'SPEED_CONTROLLED'

text list "Text list_positiveAccelStartJerkType": 40 'DIRECT'; 45 'EFFECTIVE'; 149 'USER_DEFAULT'

text list "kongding_status": 1 '状态：等待中 / 상태: 대기중'; 2 '状态：进行中 / 상태: 진행중'; 3 '状态：已完成 / 상태: 이미 완료'

text list "Text list_velocityType": 11 'CURRENT'; 40 'DIRECT'; 45 'EFFECTIVE'; 149 'USER_DEFAULT'; 312 'RESULTING'

text list "Text list_syncPositionReference": 19 'BE_SYNCHRONOUS_AT_POSITION'; 45 'EFFECTIVE'; 143 'SYNCHRONIZE_SYMMETRIC'; 144 'SYNCHRONIZE_WHEN_POSITION_REACHED'; 149 'USER_DEFAULT'

text list "Text list_move_Direction": 24 'BY_VALUE'; 45 'EFFECTIVE'; 85 'NEGATIVE'; 107 'POSITIVE'; 121 'SHORTEST_WAY'; 149 'USER_DEFAULT'

text list "Text list_negativeAccelType": 40 'DIRECT'; 45 'EFFECTIVE'; 149 'USER_DEFAULT'

text list "Text list_blendingMode": 4 'ACTIVE'; 45 'EFFECTIVE'; 61 'INACTIVE'; 149 'USER_DEFAULT'

text list "automatic_status_1": 1 '自动状态:等待 / Auto Status:Waiting / 自動状態：待機 / 자동상태:대기'; 2 '自动状态:紧急停止 / Auto Status:MergeStop / 自動状態：緊急停止 / 자동상태:비상정지'; 4 '自动状态:自动停止 / Auto Status:AtuoStop / 自動状態：自動停止 / 자동상태:자동 정지'; 8 '自动状态:出车 / Auto Status:ChuChe / 自動状態：出機 / 자동상태: 외진'; 16 '自动状态:出车到 / Auto Status:ChuCheDao / 自動状態：出機完了 / 자동상태:외진도착'; 32 '自动状态:退绕 / Auto Status:TuiRao / 自動状態：パッキング・オフ / 자동상태:언와인딩'; 64 '自动状态:卷绕 / Auto Status:JuanRao / 自動状態：巻取 / 자동상태:와인딩'; 128 '自动状态:存绕 / Auto Status:CunRao / 自動状態：逆巻取 / 자동상태:와인딩 저장'

text list "mode_enabled_1": 1 '模式:故障中 / Error / 모드: 고장중'; 2 '模式:无使能 / Disable / モード：イネーブルなし / 모드:무능력'; 4 '模式:手动 / Manual / モード：手動 / 모드:수동'; 8 '模式:定位中 / Startposition / モード：位置付け中 / 모드:위치유도'; 16 '模式:管前生头 / 모드: pipe front 스레딩'; 32 '模式:管后生头 / 모드: pipe rear 스레딩'; 64 '模式:自动 / Automatic / モード：自動 / 모드:자동'; 128 '模式:没选择 / 모드: 선택하지 않았음'; 512 '模式:生头 / モード：口付け / 모드:스레드업'

text list "Text list_Switch": 0 '已关闭'; 1 '已开启'

text list "Text list_moveTimeOutType": 169 'WITHOUT_TIME_LIMIT'; 171 'WITH_TIME_LIMIT'

text list "Text list_syncOffMode": 14 'AT_THE_END_OF_CAM_CYCLE'; 45 'EFFECTIVE'; 60 'IMMEDIATELY'; 100 'ON_MASTER_POSITION'; 101 'ON_SLAVE_POSITION'; 149 'USER_DEFAULT'

text list "KongDing_status#mig1": 0 '状态:等待中 / 상태: 대기중'; 1 '进程1:插空纱管 / 프로세스 1: 빈보빈을 삼입'; 2 '进程2:绕头 / 프로세스 2: 와인더'; 3 '进程3:罗拉送条 / 프로세스 3: 롤러 원사 공급'; 4 '进程4:锭子边卷绕 / 프로세스 4: 스핀들 사이드 와인딩'; 5 '进程5:成形弓回到原位 / 프로세스 5: 성형보우(성형호랑) 원위치 복귀'; 6 '进程6:锭子加捻 / 프로세스 6: 스핀들 연사'; 7 '进程7:牵伸、加捻 / 프로세스 7: 연신(드라프트),연사'; 8 '进程8:成形弓边至纱管底部 / 프로세스 8: 성형보우(성형호랑) 사이드에서 보빈 밑부분까지'; 9 '进程9:纱线绕几圈 / 프로세스 9: 원사를 몇바퀴 돌림'; 10 '进程10:剥掉纱管上的毛头 / 프로세스 10: 코프의 Burr 제거'; 11 '进程11:成形弓至卷绕点 / 프로세스 11: 성형보우(성형호랑)에서 와인딩 포인트까지'; 12 '进程12:进车卷绕至存绕点 / 프로세스 12: 내진 와인딩을 와인딩 저장 포인트까지 와인딩'; 13 '进程13:进车卷绕至存绕点 / 프로세스 13: 내진 와인딩을 와인딩 저장 포인트까지 와인딩'; 14 '进程14:存绕 / 프로세스 14: 와인딩 저장'

text list "mode_enabled_3": 1 '模式:故障中 / Error / 모드:고장중'; 2 '模式:无使能 / Disable / 모드:무능력'; 4 '模式:手动 / Manual / 모드:수동'; 8 '模式:定位中 / Startposition / 모드:위치유도'; 16 '模式:管前生头 / Atuomatic / 모드:pipe front 스레딩'; 32 '模式:管后生头 / NothingSelect / 모드:pipe rear 스레딩'; 64 '模式:自动 / Changing / 모드:자동'; 128 '模式:没选择 / 모드:선택하지 않았음'; 512 '模式:空锭生头 / 모드:아이들 스레드업'

text list "QainShen_Select": 2 '2段 / 2 / 2단'; 3 '3段 / 3 / 3단'

text list "Text_list_caption": 1 '自动画面 / 自動画面 / 자동화면'; 8 '手动设置 / 手動設置 / 수동설정'; 2 '手动画面 / 手動画面 / 수동화면'; 12 '张力测定 / 張力測定 / 장력 측정'; 13 '原点设置 / 原点設定 / 원점설정'; 4 '生头画面 / 生頭画面 / 스레드업화면'; 5 '报警画面 / 警報画面 / 경보화면'; 6 '保养提示 / 保全画面 / 유지보수알림'; 3 '设置画面 / 設置画面 / 설정화면'; 10 '常用调试画面 / 常用設置画面 / 상용 조정화면'; 11 '牵伸调整画面 / 연신(드라프트)조절 화면'; 14 '纱管参数设定 / 糸管パラメーター設定 / 보빈매개변수설정'; 9 '动画 / 動画 / 애니메이션'; 15 '牵伸相关 / 연신 관련'; 16 '报警记录 / 警報記録 / 경보알람기록'; 17 '参数修改画面 / パラメーター変更画面 / 매개변수 수정 화면'; 19 '配方保存画面 / レシピ保存画面 / 레시피 저장 화면'; 18 '配方选择画面 / レシピ選択画面 / 레시피선택 화면'; 7 '时间显示 / 時間表示 / 시간표시'; 20 '卷绕经验参数'; 21 '用户管理'

text list "mode_enabled_4": 1 '模式:故障中 / Error / 모드:고장중'; 2 '模式:无使能 / Disable / 모드:무능력'; 4 '模式:手动 / Manual / 모드:수동'; 8 '模式:定位中 / Startposition / 모드:위치유도'; 16 '模式:管前生头 / Atuomatic / 모드: pipe front 스레딩'; 32 '模式:管后生头 / NothingSelect / 모드: pipe rear 스레딩'; 64 '模式:自动 / Changing / 모드:자동'; 128 '模式:没选择 / 모드: 선택하지 않았음'

text list "g_i16_Calculation_0_Status": 0..6 '重新计算中'; 7 '计算完成'

graphic list "按钮": 0 '3-D red button (not pressed)_1'; 1 '3-D red button (pressed)_1'

recipe "配方_2": 总捻度 <- "ST_HMI_Var_HMI_r64NianDu_all", 支数 <- "ST_HMI_Var_HMI_r64ZhiShu_ChengSha", 牵伸捻度匹配值 <- "ST_HMI_Var_HMI_r64NianDu_QianShen_Best", 出车速度 <- "ST_HMI_Var_HMI_r64Velocity_ChuChe", 追捻开始捻度 <- "ST_HMI_Var_HMI_r64NianDu_1", 追捻锭子速度 <- "ST_HMI_Var_HMI_r64NianSu_2", 捻缩开始捻度 <- "ST_HMI_Var_HMI_r64NianDu_NianSuo", 捻缩距离 <- "ST_HMI_Var_HMI_r64Position_NianSuo", 追捻启用开关 <- "ST_HMI_Var_HMI_boNianDu_3"

recipe "配方_1": 总捻度 <- "ST_HMI_Var_HMI_r64NianDu_all", 支数 <- "ST_HMI_Var_HMI_r64ZhiShu_ChengSha", 牵伸捻度匹配值 <- "ST_HMI_Var_HMI_r64NianDu_QianShen_Best", 出车速度 <- "ST_HMI_Var_HMI_r64Velocity_ChuChe", 追捻开始捻度 <- "ST_HMI_Var_HMI_r64NianDu_1", 追捻锭子速度 <- "ST_HMI_Var_HMI_r64NianSu_2", 捻缩开始捻度 <- "ST_HMI_Var_HMI_r64NianDu_NianSuo", 捻缩距离 <- "ST_HMI_Var_HMI_r64Position_NianSuo", 追捻启用开关 <- "ST_HMI_Var_HMI_boNianDu_3"

recipe "配方_4": 总捻度 <- "ST_HMI_Var_HMI_r64NianDu_all", 支数 <- "ST_HMI_Var_HMI_r64ZhiShu_ChengSha", 牵伸捻度匹配值 <- "ST_HMI_Var_HMI_r64NianDu_QianShen_Best", 出车速度 <- "ST_HMI_Var_HMI_r64Velocity_ChuChe", 追捻开始捻度 <- "ST_HMI_Var_HMI_r64NianDu_1", 追捻锭子速度 <- "ST_HMI_Var_HMI_r64NianSu_2", 捻缩开始捻度 <- "ST_HMI_Var_HMI_r64NianDu_NianSuo", 捻缩距离 <- "ST_HMI_Var_HMI_r64Position_NianSuo", 追捻启用开关 <- "ST_HMI_Var_HMI_boNianDu_3"

recipe "配方_3": 总捻度 <- "ST_HMI_Var_HMI_r64NianDu_all", 支数 <- "ST_HMI_Var_HMI_r64ZhiShu_ChengSha", 牵伸捻度匹配值 <- "ST_HMI_Var_HMI_r64NianDu_QianShen_Best", 出车速度 <- "ST_HMI_Var_HMI_r64Velocity_ChuChe", 追捻开始捻度 <- "ST_HMI_Var_HMI_r64NianDu_1", 追捻锭子速度 <- "ST_HMI_Var_HMI_r64NianSu_2", 捻缩开始捻度 <- "ST_HMI_Var_HMI_r64NianDu_NianSuo", 捻缩距离 <- "ST_HMI_Var_HMI_r64Position_NianSuo", 追捻启用开关 <- "ST_HMI_Var_HMI_boNianDu_3"

